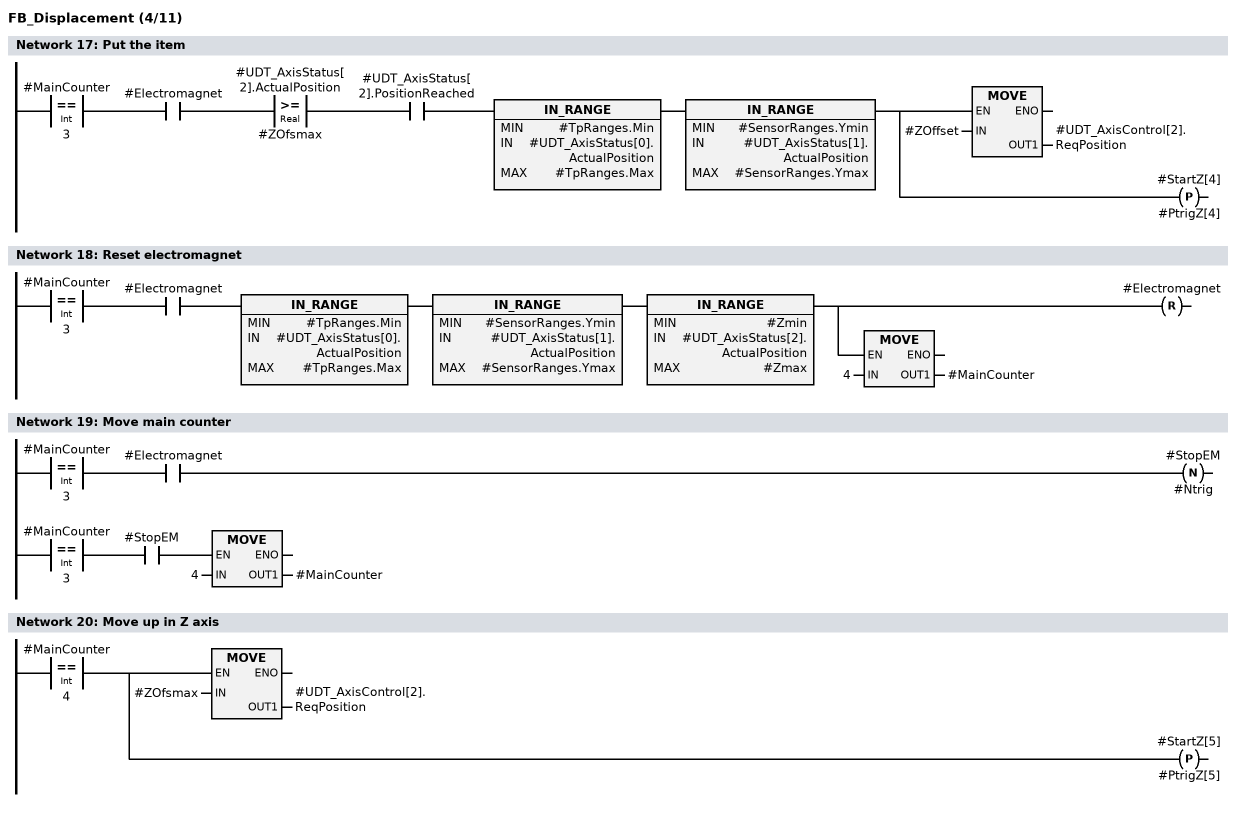
   #_w1 := (#MainCounter = 3) AND #Electromagnet AND (#UDT_AxisStatus[2].ActualPosition >= #ZOfsmax) AND #UDT_AxisStatus[2].PositionReached AND (#TpRanges.Min <= #UDT_AxisStatus[0].ActualPosition) AND (#UDT_AxisStatus[0].ActualPosition <= #TpRanges.Max) AND (#SensorRanges.Ymin <= #UDT_AxisStatus[1].ActualPosition) AND (#UDT_AxisStatus[1].ActualPosition <= #SensorRanges.Ymax);
   IF #_w1 THEN #UDT_AxisControl[2].ReqPosition := #ZOffset; END_IF;
   #StartZ[4] := #_w1 AND NOT #PtrigZ[4];   // rising edge
   #PtrigZ[4] := #_w1;
END_REGION

REGION Network 18: Reset electromagnet
   RUNG wire#powerrail
      { S7_Templates := "SrcType := Int" } EQ_Contact(in1 := #MainCounter, in2 := 3)
      Contact( #Electromagnet )
      { S7_Templates := "SrcType := Real" } InRange(min := #TpRanges.Min, in := #UDT_AxisStatus[0].ActualPosition, max := #TpRanges.Max)
      { S7_Templates := "SrcType := Real" } InRange(min := #SensorRanges.Ymin, in := #UDT_AxisStatus[1].ActualPosition, max := #SensorRanges.Ymax)
      { S7_Templates := "SrcType := Real" } InRange(min := #Zmin, in := #UDT_AxisStatus[2].ActualPosition, max := #Zmax)
      wire#w1
      R_Coil( #Electromagnet )
   END_RUNG
   RUNG wire#w1
      Move(in := 4, out1 => #MainCounter)
   END_RUNG
   // the same network as SCL:
   #_w1 := (#MainCounter = 3) AND #Electromagnet AND (#TpRanges.Min <= #UDT_AxisStatus[0].ActualPosition) AND (#UDT_AxisStatus[0].ActualPosition <= #TpRanges.Max) AND (#SensorRanges.Ymin <= #UDT_AxisStatus[1].ActualPosition) AND (#UDT_AxisStatus[1].ActualPosition <= #SensorRanges.Ymax) AND (#Zmin <= #UDT_AxisStatus[2].ActualPosition) AND (#UDT_AxisStatus[2].ActualPosition <= #Zmax);
   IF #_w1 THEN
       #Electromagnet := FALSE;
       #MainCounter := 4;
   END_IF;
END_REGION

REGION Network 19: Move main counter
   #_w1 := (#MainCounter = 3) AND #Electromagnet;
   #StopEM := NOT #_w1 AND #Ntrig;   // falling edge
   #Ntrig := #_w1;
   IF (#MainCounter = 3) AND #StopEM THEN #MainCounter := 4; END_IF;
END_REGION

REGION Network 20: Move up in Z axis
   #_w1 := #MainCounter = 4;
   IF #_w1 THEN #UDT_AxisControl[2].ReqPosition := #ZOfsmax; END_IF;
   #StartZ[5] := #_w1 AND NOT #PtrigZ[5];   // rising edge
   #PtrigZ[5] := #_w1;
END_REGION

REGION Network 21: Move to the previous or starting position
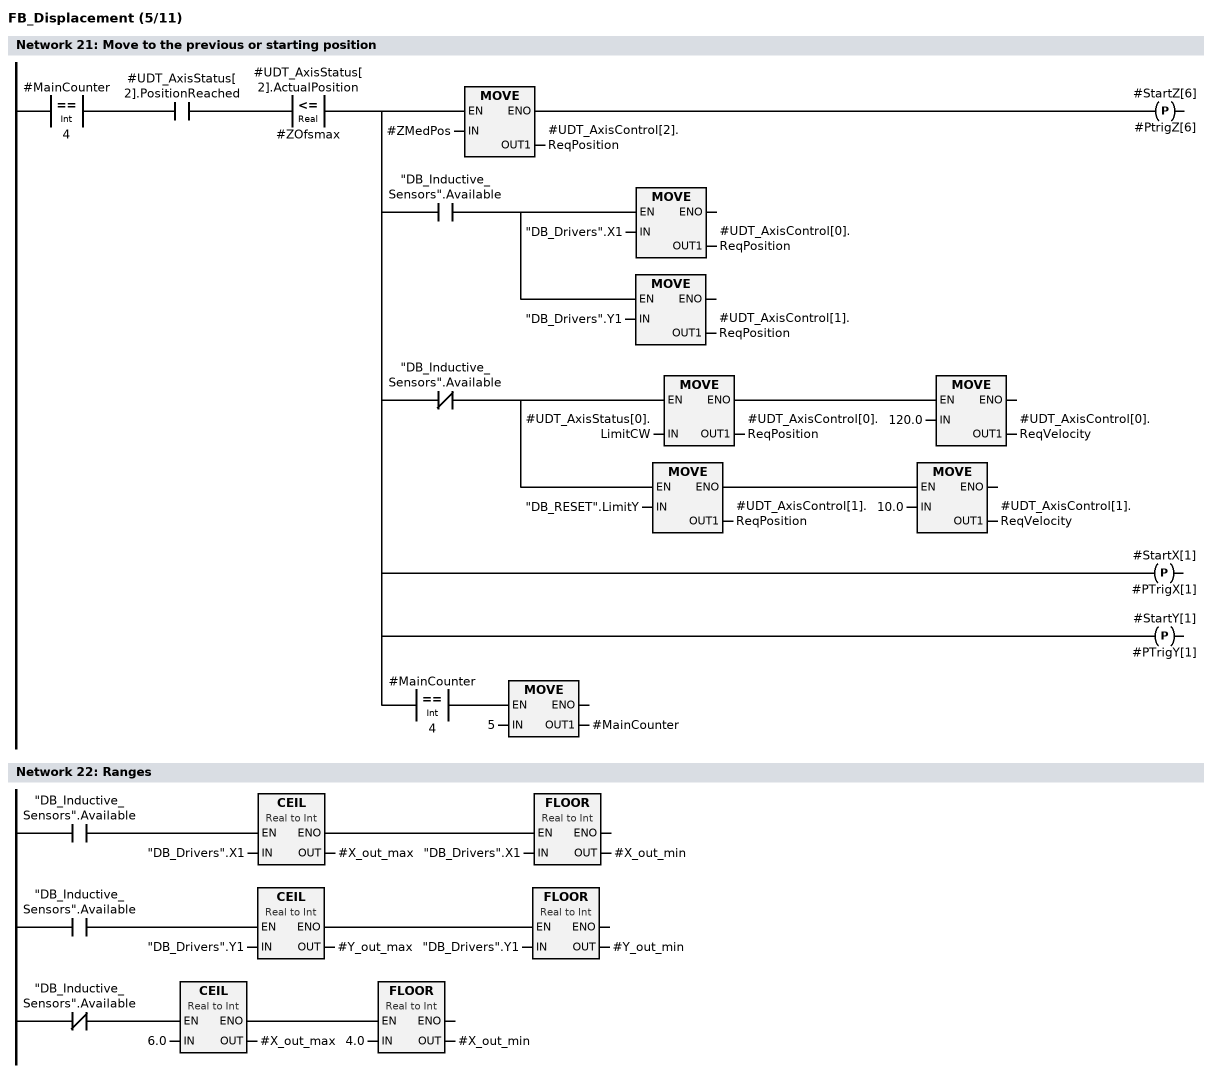
   #_w1 := (#MainCounter = 4) AND #UDT_AxisStatus[2].PositionReached AND (#UDT_AxisStatus[2].ActualPosition <= #ZOfsmax);
   IF #_w1 THEN #UDT_AxisControl[2].ReqPosition := #ZMedPos; END_IF;
   #StartZ[6] := #_w1 AND NOT #PtrigZ[6];   // rising edge
   #PtrigZ[6] := #_w1;
   IF #_w1 AND "DB_Inductive_Sensors".Available THEN
       #UDT_AxisControl[0].ReqPosition := "DB_Drivers".X1;
       #UDT_AxisControl[1].ReqPosition := "DB_Drivers".Y1;
   END_IF;
   IF #_w1 AND NOT "DB_Inductive_Sensors".Available THEN
       #UDT_AxisControl[0].ReqPosition := #UDT_AxisStatus[0].LimitCW;
       #UDT_AxisControl[0].ReqVelocity := 120.0;
       #UDT_AxisControl[1].ReqPosition := "DB_RESET".LimitY;
       #UDT_AxisControl[1].ReqVelocity := 10.0;
   END_IF;
   #StartX[1] := #_w1 AND NOT #PTrigX[1];   // rising edge
   #PTrigX[1] := #_w1;
   #StartY[1] := #_w1 AND NOT #PTrigY[1];   // rising edge
   #PTrigY[1] := #_w1;
   IF #_w1 AND (#MainCounter = 4) THEN #MainCounter := 5; END_IF;
END_REGION

REGION Network 22: Ranges
   IF "DB_Inductive_Sensors".Available THEN
       #X_out_max := CEIL("DB_Drivers".X1);
       #X_out_min := FLOOR("DB_Drivers".X1);
       #Y_out_max := CEIL("DB_Drivers".Y1);
       #Y_out_min := FLOOR("DB_Drivers".Y1);
   END_IF;
   IF NOT "DB_Inductive_Sensors".Available THEN
       #X_out_max := CEIL(6.0);
       #X_out_min := FLOOR(4.0);
   END_IF;
END_REGION

REGION Network 23: Places occupied
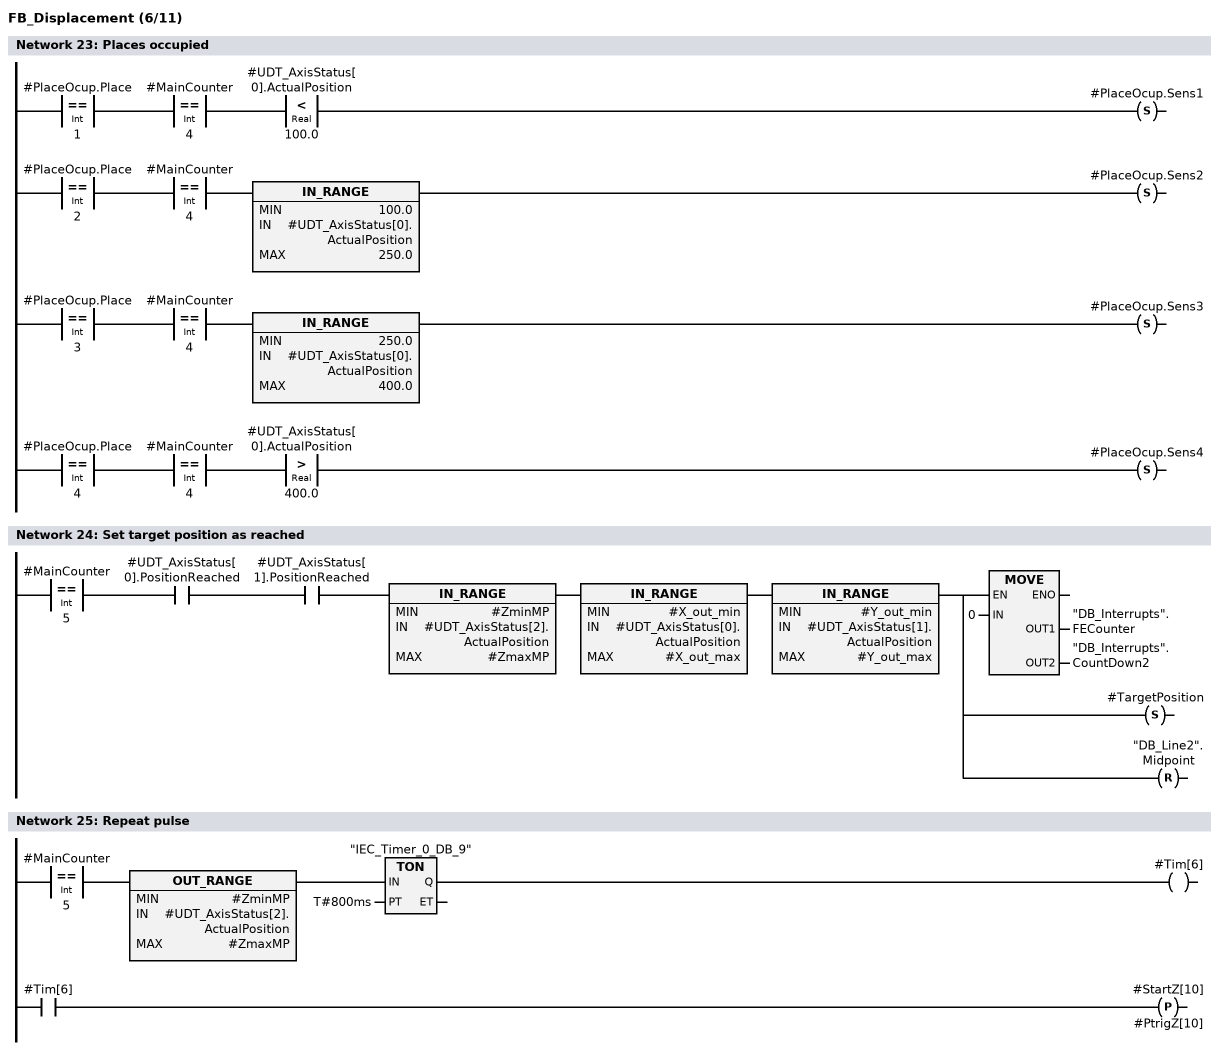
   RUNG wire#powerrail
      { S7_Templates := "SrcType := Int" } EQ_Contact(in1 := #PlaceOcup.Place, in2 := 1)
      { S7_Templates := "SrcType := Int" } EQ_Contact(in1 := #MainCounter, in2 := 4)
      { S7_Templates := "SrcType := Real" } LT_Contact(in1 := #UDT_AxisStatus[0].ActualPosition, in2 := 100.0)
      S_Coil( #PlaceOcup.Sens1 )
   END_RUNG
   RUNG wire#powerrail
      { S7_Templates := "SrcType := Int" } EQ_Contact(in1 := #PlaceOcup.Place, in2 := 2)
      { S7_Templates := "SrcType := Int" } EQ_Contact(in1 := #MainCounter, in2 := 4)
      { S7_Templates := "SrcType := Real" } InRange(min := 100.0, in := #UDT_AxisStatus[0].ActualPosition, max := 250.0)
      S_Coil( #PlaceOcup.Sens2 )
   END_RUNG
   RUNG wire#powerrail
      { S7_Templates := "SrcType := Int" } EQ_Contact(in1 := #PlaceOcup.Place, in2 := 3)
      { S7_Templates := "SrcType := Int" } EQ_Contact(in1 := #MainCounter, in2 := 4)
      { S7_Templates := "SrcType := Real" } InRange(min := 250.0, in := #UDT_AxisStatus[0].ActualPosition, max := 400.0)
      S_Coil( #PlaceOcup.Sens3 )
   END_RUNG
   RUNG wire#powerrail
      { S7_Templates := "SrcType := Int" } EQ_Contact(in1 := #PlaceOcup.Place, in2 := 4)
      { S7_Templates := "SrcType := Int" } EQ_Contact(in1 := #MainCounter, in2 := 4)
      { S7_Templates := "SrcType := Real" } GT_Contact(in1 := #UDT_AxisStatus[0].ActualPosition, in2 := 400.0)
      S_Coil( #PlaceOcup.Sens4 )
   END_RUNG
   // the same network as SCL:
   IF (#PlaceOcup.Place = 1) AND (#MainCounter = 4) AND (#UDT_AxisStatus[0].ActualPosition < 100.0) THEN
       #PlaceOcup.Sens1 := TRUE;
   END_IF;
   IF (#PlaceOcup.Place = 2) AND (#MainCounter = 4) AND (100.0 <= #UDT_AxisStatus[0].ActualPosition) AND (#UDT_AxisStatus[0].ActualPosition <= 250.0) THEN
       #PlaceOcup.Sens2 := TRUE;
   END_IF;
   IF (#PlaceOcup.Place = 3) AND (#MainCounter = 4) AND (250.0 <= #UDT_AxisStatus[0].ActualPosition) AND (#UDT_AxisStatus[0].ActualPosition <= 400.0) THEN
       #PlaceOcup.Sens3 := TRUE;
   END_IF;
   IF (#PlaceOcup.Place = 4) AND (#MainCounter = 4) AND (#UDT_AxisStatus[0].ActualPosition > 400.0) THEN
       #PlaceOcup.Sens4 := TRUE;
   END_IF;
END_REGION

REGION Network 24: Set target position as reached
   RUNG wire#powerrail
      { S7_Templates := "SrcType := Int" } EQ_Contact(in1 := #MainCounter, in2 := 5)
      Contact( #UDT_AxisStatus[0].PositionReached )
      Contact( #UDT_AxisStatus[1].PositionReached )
      { S7_Templates := "SrcType := Real" } InRange(min := #ZminMP, in := #UDT_AxisStatus[2].ActualPosition, max := #ZmaxMP)
      { S7_Templates := "SrcType := Real" } InRange(min := #X_out_min, in := #UDT_AxisStatus[0].ActualPosition, max := #X_out_max)
      { S7_Templates := "SrcType := Real" } InRange(min := #Y_out_min, in := #UDT_AxisStatus[1].ActualPosition, max := #Y_out_max)
      wire#w1
      Move(in := 0, out1 => "DB_Interrupts".FECounter, out2 => "DB_Interrupts".CountDown2)
   END_RUNG
   RUNG wire#w1
      S_Coil( #TargetPosition )
   END_RUNG
   RUNG wire#w1
      R_Coil( "DB_Line2".Midpoint )
   END_RUNG
   // the same network as SCL:
   IF (#MainCounter = 5) AND #UDT_AxisStatus[0].PositionReached AND #UDT_AxisStatus[1].PositionReached AND (#ZminMP <= #UDT_AxisStatus[2].ActualPosition) AND (#UDT_AxisStatus[2].ActualPosition <= #ZmaxMP) AND (#X_out_min <= #UDT_AxisStatus[0].ActualPosition) AND (#UDT_AxisStatus[0].ActualPosition <= #X_out_max) AND (#Y_out_min <= #UDT_AxisStatus[1].ActualPosition) AND (#UDT_AxisStatus[1].ActualPosition <= #Y_out_max) THEN
       "DB_Interrupts".FECounter := 0;
       "DB_Interrupts".CountDown2 := 0;
       #TargetPosition := TRUE;
       "DB_Line2".Midpoint := FALSE;
   END_IF;
END_REGION

REGION Network 25: Repeat pulse
   "IEC_Timer_0_DB_9".TON(IN := (#MainCounter = 5) AND ((#UDT_AxisStatus[2].ActualPosition < #ZminMP) OR (#UDT_AxisStatus[2].ActualPosition > #ZmaxMP)),
                          PT := T#800ms);
   #Tim[6] := "IEC_Timer_0_DB_9".Q;
   #StartZ[10] := #Tim[6] AND NOT #PtrigZ[10];   // rising edge
   #PtrigZ[10] := #Tim[6];
END_REGION

REGION Network 26: Additional timers
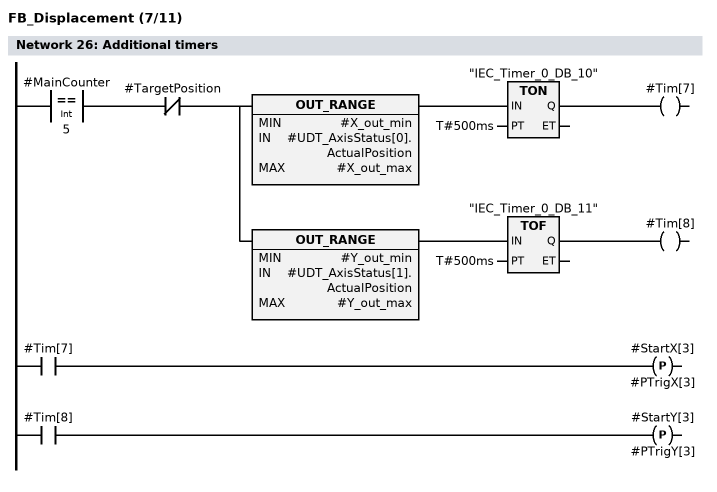
   #_w1 := (#MainCounter = 5) AND NOT #TargetPosition;
   "IEC_Timer_0_DB_10".TON(IN := #_w1 AND ((#UDT_AxisStatus[0].ActualPosition < #X_out_min) OR (#UDT_AxisStatus[0].ActualPosition > #X_out_max)),
                           PT := T#500ms);
   #Tim[7] := "IEC_Timer_0_DB_10".Q;
   "IEC_Timer_0_DB_11".TOF(IN := #_w1 AND ((#UDT_AxisStatus[1].ActualPosition < #Y_out_min) OR (#UDT_AxisStatus[1].ActualPosition > #Y_out_max)),
                           PT := T#500ms);
   #Tim[8] := "IEC_Timer_0_DB_11".Q;
   #StartX[3] := #Tim[7] AND NOT #PTrigX[3];   // rising edge
   #PTrigX[3] := #Tim[7];
   #StartY[3] := #Tim[8] AND NOT #PTrigY[3];   // rising edge
   #PTrigY[3] := #Tim[8];
END_REGION

REGION Network 27: Item was detected. Interrupt is active.
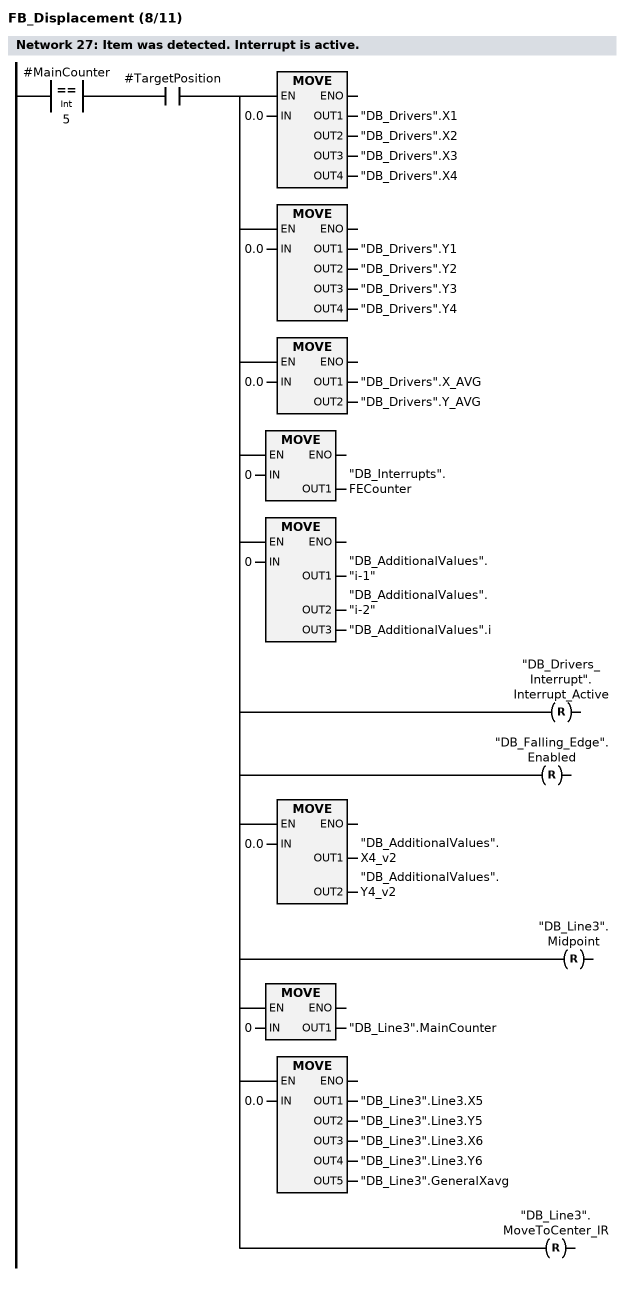
   RUNG wire#powerrail
      { S7_Templates := "SrcType := Int" } EQ_Contact(in1 := #MainCounter, in2 := 5)
      Contact( #TargetPosition )
      wire#w1
      Move(in := 0.0, out1 => "DB_Drivers".X1, out2 => "DB_Drivers".X2, out3 => "DB_Drivers".X3, out4 => "DB_Drivers".X4)
   END_RUNG
   RUNG wire#w1
      Move(in := 0.0, out1 => "DB_Drivers".Y1, out2 => "DB_Drivers".Y2, out3 => "DB_Drivers".Y3, out4 => "DB_Drivers".Y4)
   END_RUNG
   RUNG wire#w1
      Move(in := 0.0, out1 => "DB_Drivers".X_AVG, out2 => "DB_Drivers".Y_AVG)
   END_RUNG
   RUNG wire#w1
      Move(in := 0, out1 => "DB_Interrupts".FECounter)
   END_RUNG
   RUNG wire#w1
      Move(in := 0, out1 => "DB_AdditionalValues"."i-1", out2 => "DB_AdditionalValues"."i-2", out3 => "DB_AdditionalValues".i)
   END_RUNG
   RUNG wire#w1
      R_Coil( "DB_Drivers_Interrupt".Interrupt_Active )
   END_RUNG
   RUNG wire#w1
      R_Coil( "DB_Falling_Edge".Enabled )
   END_RUNG
   RUNG wire#w1
      Move(in := 0.0, out1 => "DB_AdditionalValues".X4_v2, out2 => "DB_AdditionalValues".Y4_v2)
   END_RUNG
   RUNG wire#w1
      R_Coil( "DB_Line3".Midpoint )
   END_RUNG
   RUNG wire#w1
      Move(in := 0, out1 => "DB_Line3".MainCounter)
   END_RUNG
   RUNG wire#w1
      Move(in := 0.0, out1 => "DB_Line3".Line3.X5, out2 => "DB_Line3".Line3.Y5, out3 => "DB_Line3".Line3.X6, out4 => "DB_Line3".Line3.Y6, out5 => "DB_Line3".GeneralXavg)
   END_RUNG
   RUNG wire#w1
      R_Coil( "DB_Line3".MoveToCenter_IR )
   END_RUNG
   // the same network as SCL:
   IF (#MainCounter = 5) AND #TargetPosition THEN
       "DB_Drivers".X1 := 0.0;
       "DB_Drivers".X2 := 0.0;
       "DB_Drivers".X3 := 0.0;
       "DB_Drivers".X4 := 0.0;
       "DB_Drivers".Y1 := 0.0;
       "DB_Drivers".Y2 := 0.0;
       "DB_Drivers".Y3 := 0.0;
       "DB_Drivers".Y4 := 0.0;
       "DB_Drivers".X_AVG := 0.0;
       "DB_Drivers".Y_AVG := 0.0;
       "DB_Interrupts".FECounter := 0;
       "DB_AdditionalValues"."i-1" := 0;
       "DB_AdditionalValues"."i-2" := 0;
       "DB_AdditionalValues".i := 0;
       "DB_Drivers_Interrupt".Interrupt_Active := FALSE;
       "DB_Falling_Edge".Enabled := FALSE;
       "DB_AdditionalValues".X4_v2 := 0.0;
       "DB_AdditionalValues".Y4_v2 := 0.0;
       "DB_Line3".Midpoint := FALSE;
       "DB_Line3".MainCounter := 0;
       "DB_Line3".Line3.X5 := 0.0;
       "DB_Line3".Line3.Y5 := 0.0;
       "DB_Line3".Line3.X6 := 0.0;
       "DB_Line3".Line3.Y6 := 0.0;
       "DB_Line3".GeneralXavg := 0.0;
       "DB_Line3".MoveToCenter_IR := FALSE;
   END_IF;
END_REGION

REGION Network 28: Start Movement Command in X axis
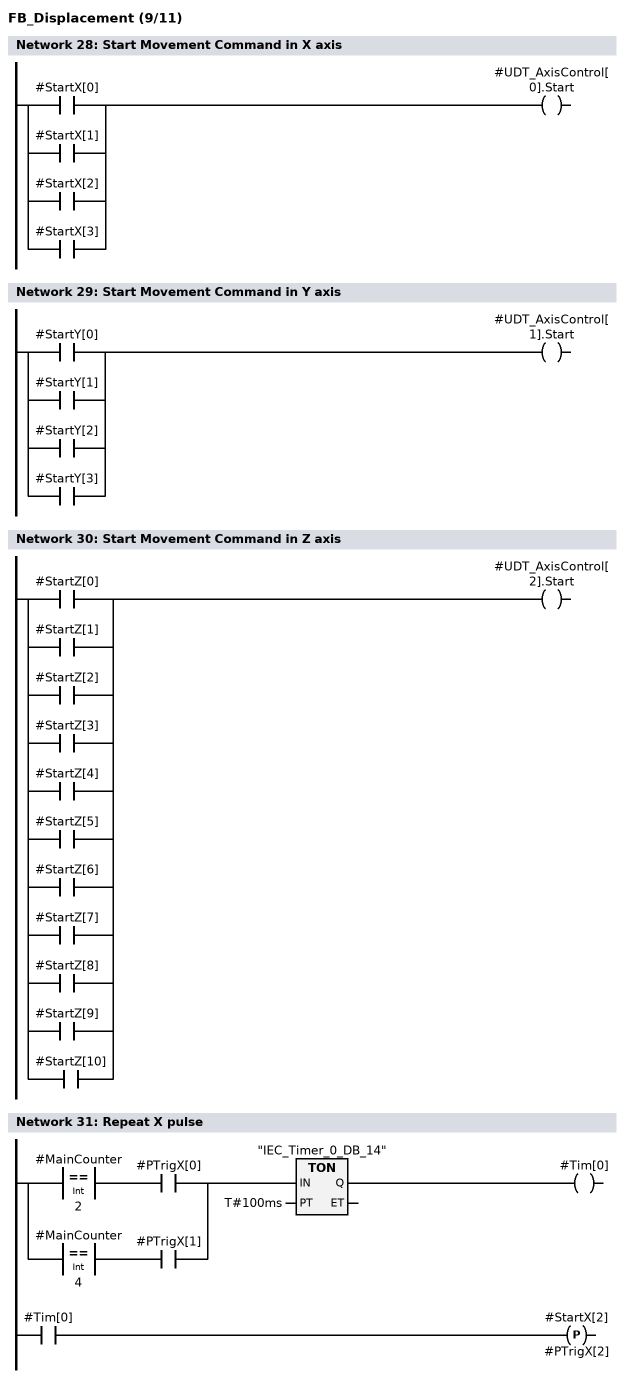
   RUNG wire#powerrail
      Contact( #StartX[0] )
      wire#w1
      Coil( #UDT_AxisControl[0].Start )
   END_RUNG
   RUNG wire#powerrail
      Contact( #StartX[1] )
   END_RUNG wire#w1
   RUNG wire#powerrail
      Contact( #StartX[2] )
   END_RUNG wire#w1
   RUNG wire#powerrail
      Contact( #StartX[3] )
   END_RUNG wire#w1
   // the same network as SCL:
   #UDT_AxisControl[0].Start := #StartX[0] OR #StartX[1] OR #StartX[2] OR #StartX[3];
END_REGION

REGION Network 29: Start Movement Command in Y axis
   RUNG wire#powerrail
      Contact( #StartY[0] )
      wire#w1
      Coil( #UDT_AxisControl[1].Start )
   END_RUNG
   RUNG wire#powerrail
      Contact( #StartY[1] )
   END_RUNG wire#w1
   RUNG wire#powerrail
      Contact( #StartY[2] )
   END_RUNG wire#w1
   RUNG wire#powerrail
      Contact( #StartY[3] )
   END_RUNG wire#w1
   // the same network as SCL:
   #UDT_AxisControl[1].Start := #StartY[0] OR #StartY[1] OR #StartY[2] OR #StartY[3];
END_REGION

REGION Network 30: Start Movement Command in Z axis
   RUNG wire#powerrail
      Contact( #StartZ[0] )
      wire#w1
      Coil( #UDT_AxisControl[2].Start )
   END_RUNG
   RUNG wire#powerrail
      Contact( #StartZ[1] )
   END_RUNG wire#w1
   RUNG wire#powerrail
      Contact( #StartZ[2] )
   END_RUNG wire#w1
   RUNG wire#powerrail
      Contact( #StartZ[3] )
   END_RUNG wire#w1
   RUNG wire#powerrail
      Contact( #StartZ[4] )
   END_RUNG wire#w1
   RUNG wire#powerrail
      Contact( #StartZ[5] )
   END_RUNG wire#w1
   RUNG wire#powerrail
      Contact( #StartZ[6] )
   END_RUNG wire#w1
   RUNG wire#powerrail
      Contact( #StartZ[7] )
   END_RUNG wire#w1
   RUNG wire#powerrail
      Contact( #StartZ[8] )
   END_RUNG wire#w1
   RUNG wire#powerrail
      Contact( #StartZ[9] )
   END_RUNG wire#w1
   RUNG wire#powerrail
      Contact( #StartZ[10] )
   END_RUNG wire#w1
   // the same network as SCL:
   #UDT_AxisControl[2].Start := #StartZ[0] OR #StartZ[1] OR #StartZ[2] OR #StartZ[3] OR #StartZ[4] OR #StartZ[5] OR #StartZ[6] OR #StartZ[7] OR #StartZ[8] OR #StartZ[9] OR #StartZ[10];
END_REGION

REGION Network 31: Repeat X pulse
   "IEC_Timer_0_DB_14".TON(IN := ((#MainCounter = 2) AND #PTrigX[0]) OR ((#MainCounter = 4) AND #PTrigX[1]),
                           PT := T#100ms);
   #Tim[0] := "IEC_Timer_0_DB_14".Q;
   #StartX[2] := #Tim[0] AND NOT #PTrigX[2];   // rising edge
   #PTrigX[2] := #Tim[0];
END_REGION

REGION Network 32: Repeat Y pulse
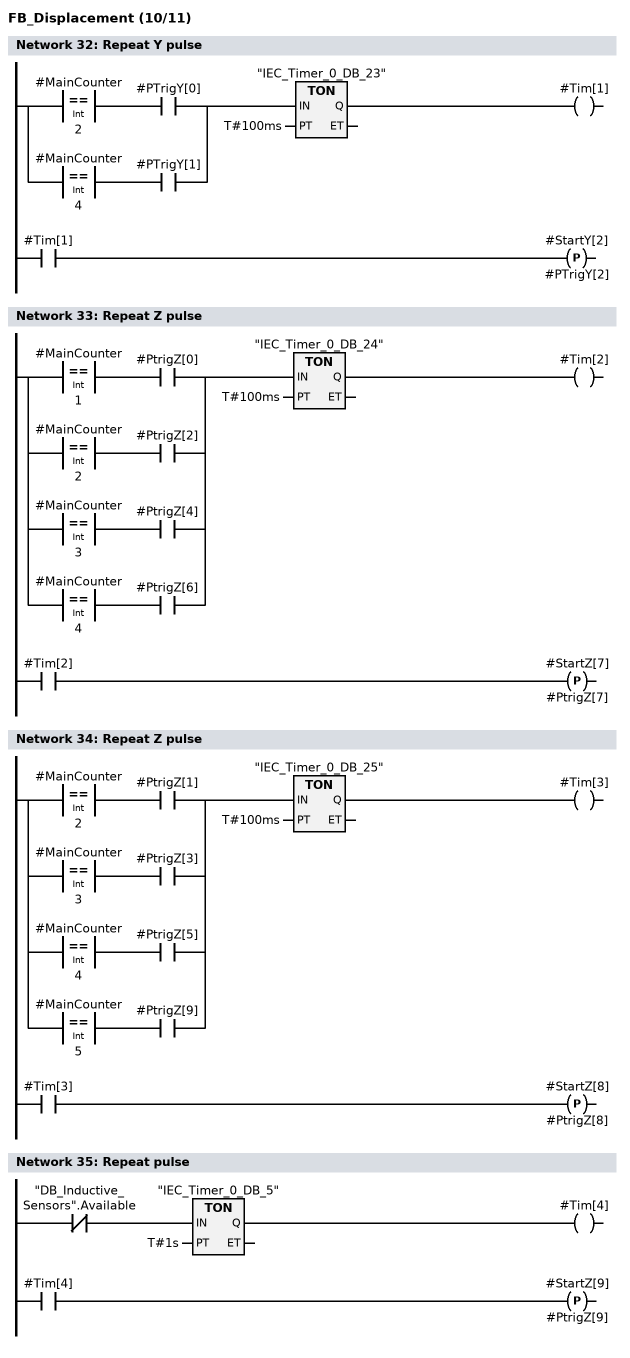
   "IEC_Timer_0_DB_23".TON(IN := ((#MainCounter = 2) AND #PTrigY[0]) OR ((#MainCounter = 4) AND #PTrigY[1]),
                           PT := T#100ms);
   #Tim[1] := "IEC_Timer_0_DB_23".Q;
   #StartY[2] := #Tim[1] AND NOT #PTrigY[2];   // rising edge
   #PTrigY[2] := #Tim[1];
END_REGION

REGION Network 33: Repeat Z pulse
   "IEC_Timer_0_DB_24".TON(IN := ((#MainCounter = 1) AND #PtrigZ[0]) OR ((#MainCounter = 2) AND #PtrigZ[2]) OR ((#MainCounter = 3) AND #PtrigZ[4]) OR ((#MainCounter = 4) AND #PtrigZ[6]),
                           PT := T#100ms);
   #Tim[2] := "IEC_Timer_0_DB_24".Q;
   #StartZ[7] := #Tim[2] AND NOT #PtrigZ[7];   // rising edge
   #PtrigZ[7] := #Tim[2];
END_REGION

REGION Network 34: Repeat Z pulse
   "IEC_Timer_0_DB_25".TON(IN := ((#MainCounter = 2) AND #PtrigZ[1]) OR ((#MainCounter = 3) AND #PtrigZ[3]) OR ((#MainCounter = 4) AND #PtrigZ[5]) OR ((#MainCounter = 5) AND #PtrigZ[9]),
                           PT := T#100ms);
   #Tim[3] := "IEC_Timer_0_DB_25".Q;
   #StartZ[8] := #Tim[3] AND NOT #PtrigZ[8];   // rising edge
   #PtrigZ[8] := #Tim[3];
END_REGION

REGION Network 35: Repeat pulse
   "IEC_Timer_0_DB_5".TON(IN := NOT "DB_Inductive_Sensors".Available, PT := T#1s);
   #Tim[4] := "IEC_Timer_0_DB_5".Q;
   #StartZ[9] := #Tim[4] AND NOT #PtrigZ[9];   // rising edge
   #PtrigZ[9] := #Tim[4];
END_REGION

REGION Network 36
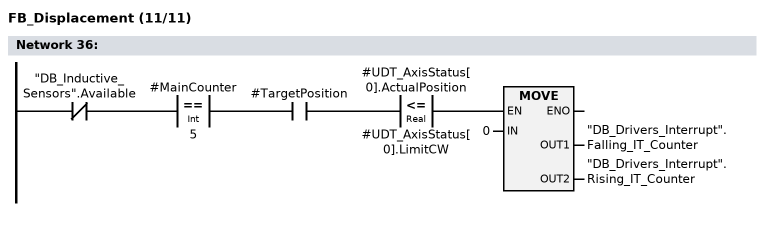
   RUNG wire#powerrail
      I_Contact( "DB_Inductive_Sensors".Available )
      { S7_Templates := "SrcType := Int" } EQ_Contact(in1 := #MainCounter, in2 := 5)
      Contact( #TargetPosition )
      { S7_Templates := "SrcType := Real" } LE_Contact(in1 := #UDT_AxisStatus[0].ActualPosition, in2 := #UDT_AxisStatus[0].LimitCW)
      Move(in := 0, out1 => "DB_Drivers_Interrupt".Falling_IT_Counter, out2 => "DB_Drivers_Interrupt".Rising_IT_Counter)
   END_RUNG
   // the same network as SCL:
   IF NOT "DB_Inductive_Sensors".Available AND (#MainCounter = 5) AND #TargetPosition AND (#UDT_AxisStatus[0].ActualPosition <= #UDT_AxisStatus[0].LimitCW) THEN
       "DB_Drivers_Interrupt".Falling_IT_Counter := 0;
       "DB_Drivers_Interrupt".Rising_IT_Counter := 0;
   END_IF;
END_REGION
END_FUNCTION_BLOCK

// folder: Displacement/Object displacement/Inductive Sensors

FUNCTION_BLOCK "FB_Inductive_Sensors"   // FB14, LAD
{ S7_Optimized_Access := 'TRUE' }
VERSION : 0.1
   VAR_INPUT
      Sensor_1 : Bool;
      Sensor_2 : Bool;
      Sensor_3 : Bool;
      Sensor_4 : Bool;
   END_VAR
   VAR_OUTPUT
      Available : Bool;
      "Sensor CO" : Struct   // Numbers and coordinates of the first available sensor
         Sensor_Pos_X : Real;
         Sensor_Pos_Y : Real;
         SensorNumber : Int;
      END_STRUCT;
      "Sensor CO Reach" : Struct   // Ranges of each sensors
         "X min" : Real;
         "X max" : Real;
         "Y min" : Real;
         "Y max" : Real;
      END_STRUCT;
   END_VAR
   VAR
      "Ind Sensor_CO" : Struct   // Numbers and coordinates of each sensor
         "Sensor 1" : Struct
            "Pos X" : Real := 23.0;   // 23 mm
            "Pos Y" : Real := 284.0;   // 284
            SensorNumber : Int;
         END_STRUCT;
         "Sensor 2" : Struct
            "Pos X" : Real := 167.0;   // 167 mm
            "Pos Y" : Real := 284.0;
            SensorNumber : Int;
         END_STRUCT;
         "Sensor 3" : Struct
            "Pos X" : Real := 313.0;   // 313 mm
            "Pos Y" : Real := 284.0;
            SensorNumber : Int;
         END_STRUCT;
         "Sensor 4" : Struct
            "Pos X" : Real := 463.0;   // 463 mm
            "Pos Y" : Real := 284.0;
            SensorNumber : Int;
         END_STRUCT;
      END_STRUCT;
      "Limit Y" : Real;
   END_VAR
BEGIN

REGION Network 1: Inductive Sensors
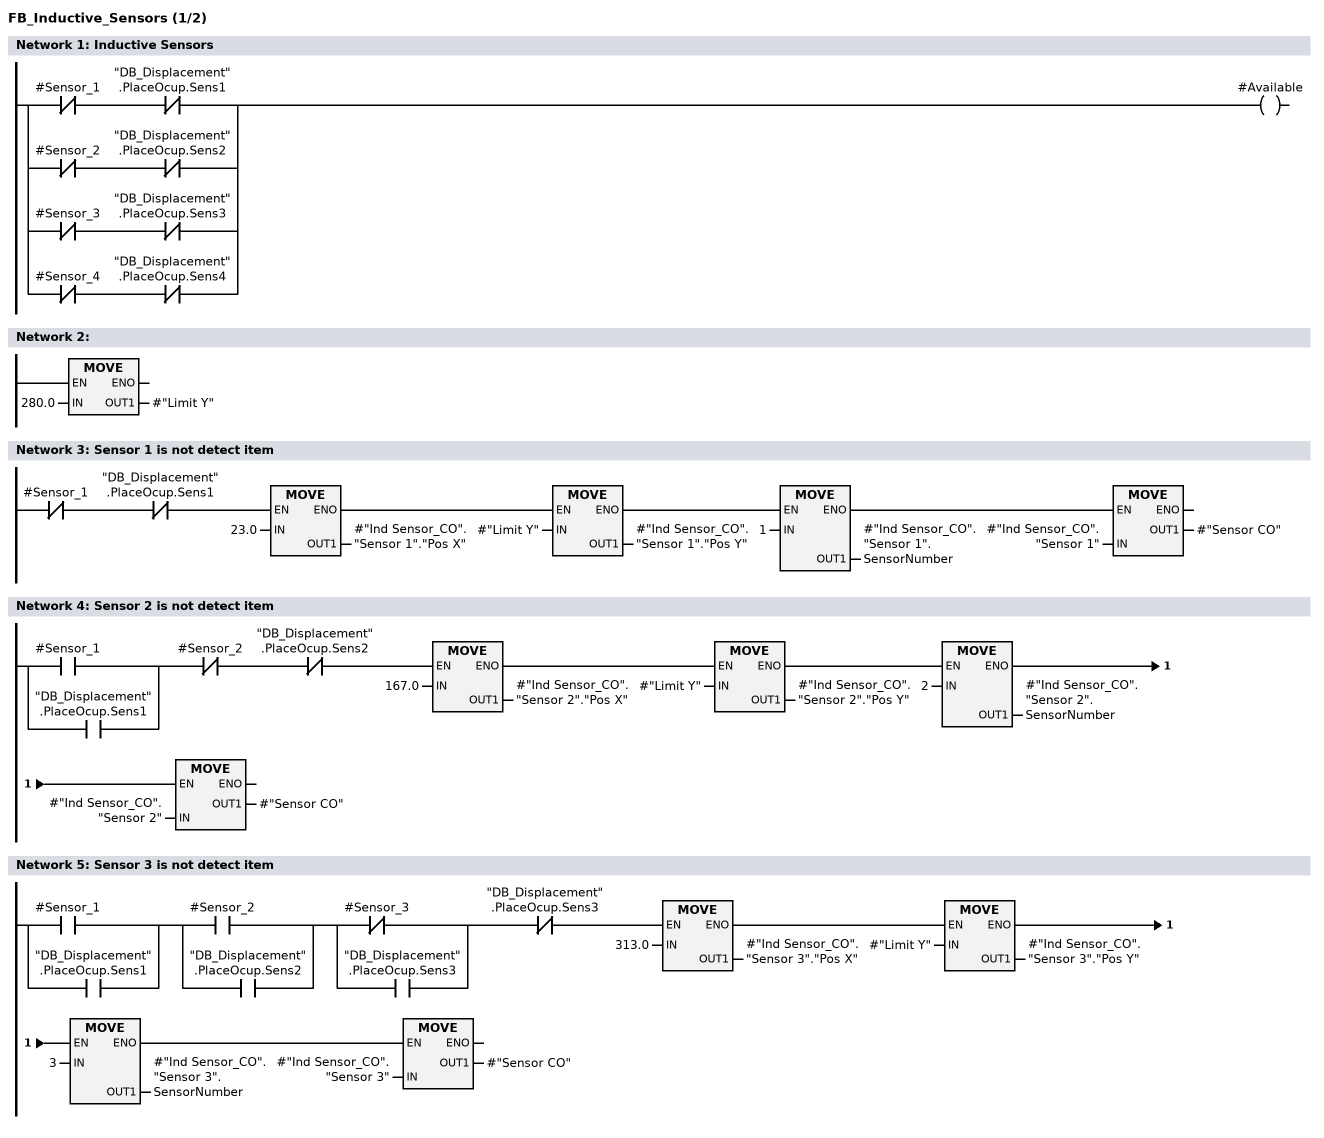
   RUNG wire#powerrail
      I_Contact( #Sensor_1 )
      I_Contact( "DB_Displacement".PlaceOcup.Sens1 )
      wire#w1
      Coil( #Available )
   END_RUNG
   RUNG wire#powerrail
      I_Contact( #Sensor_2 )
      I_Contact( "DB_Displacement".PlaceOcup.Sens2 )
   END_RUNG wire#w1